       "CompALTA-MTA".Static_60 := 2;
   END_IF;
END_REGION

REGION Network 12
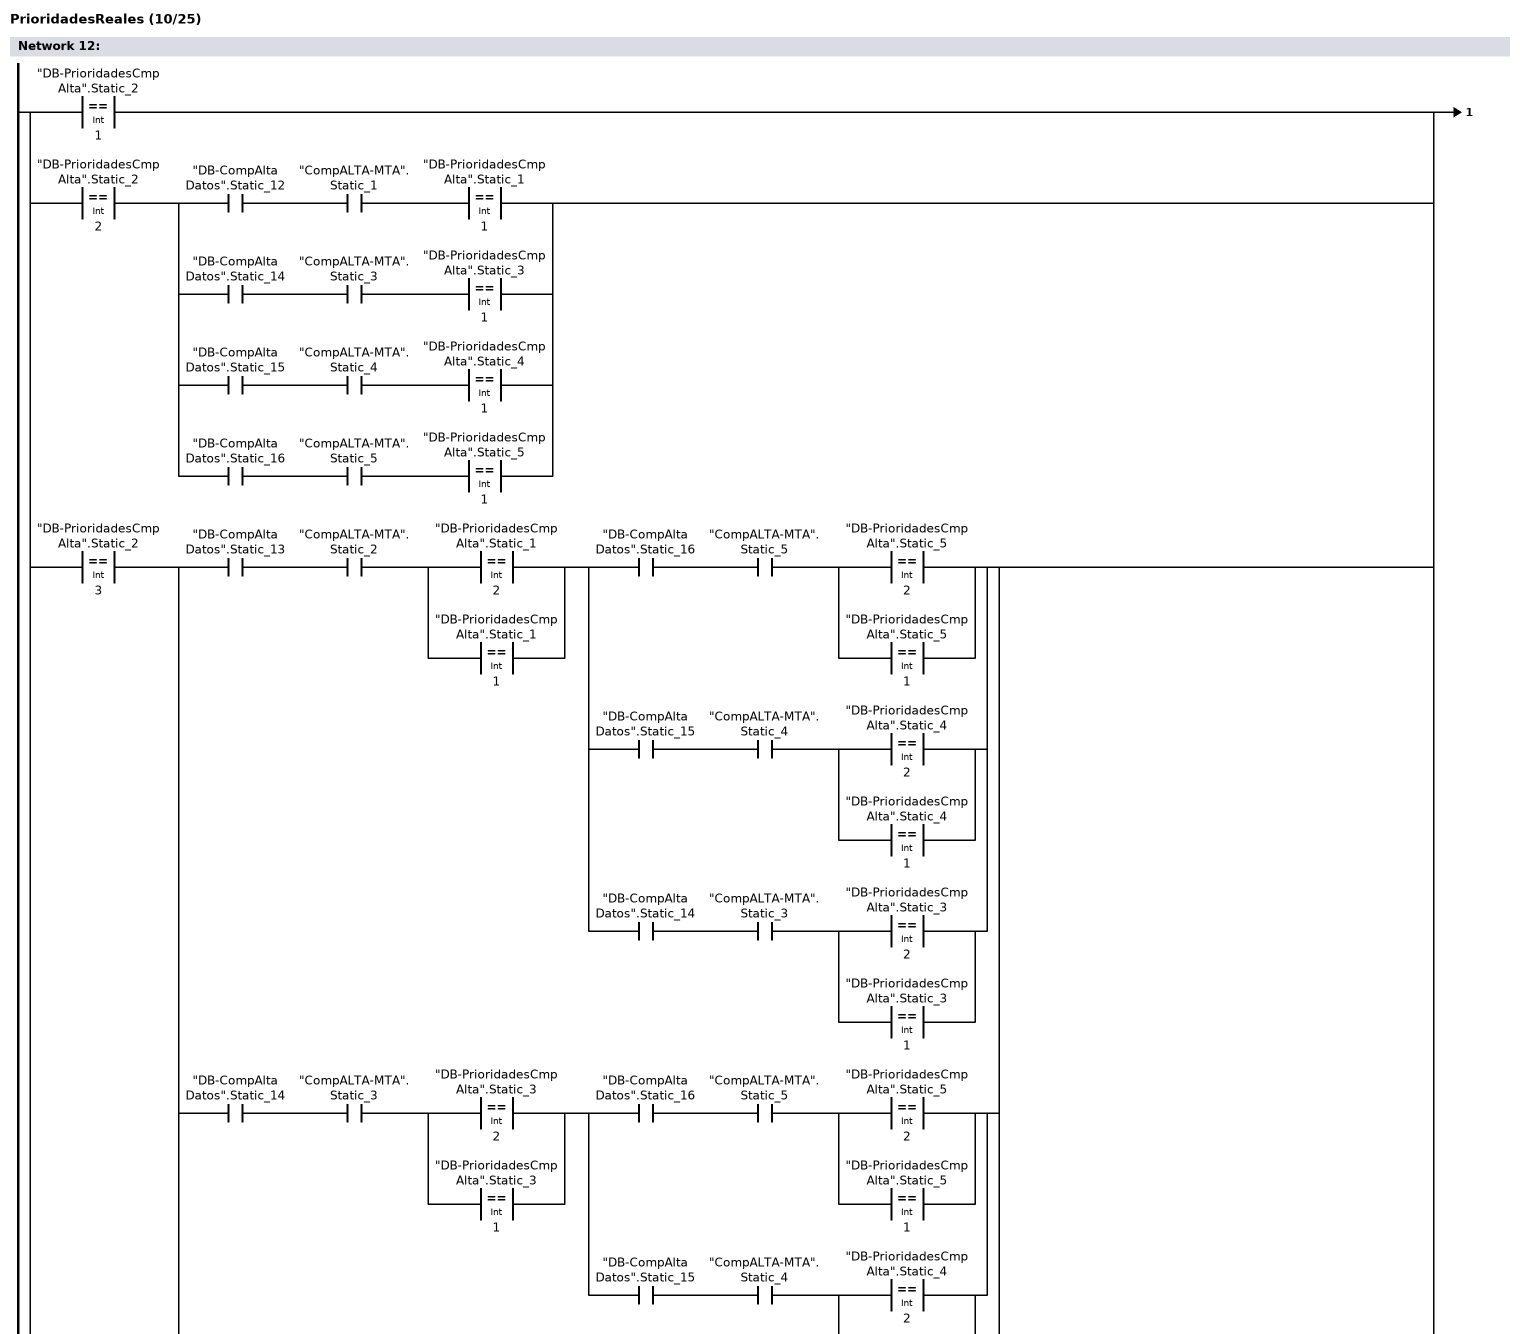
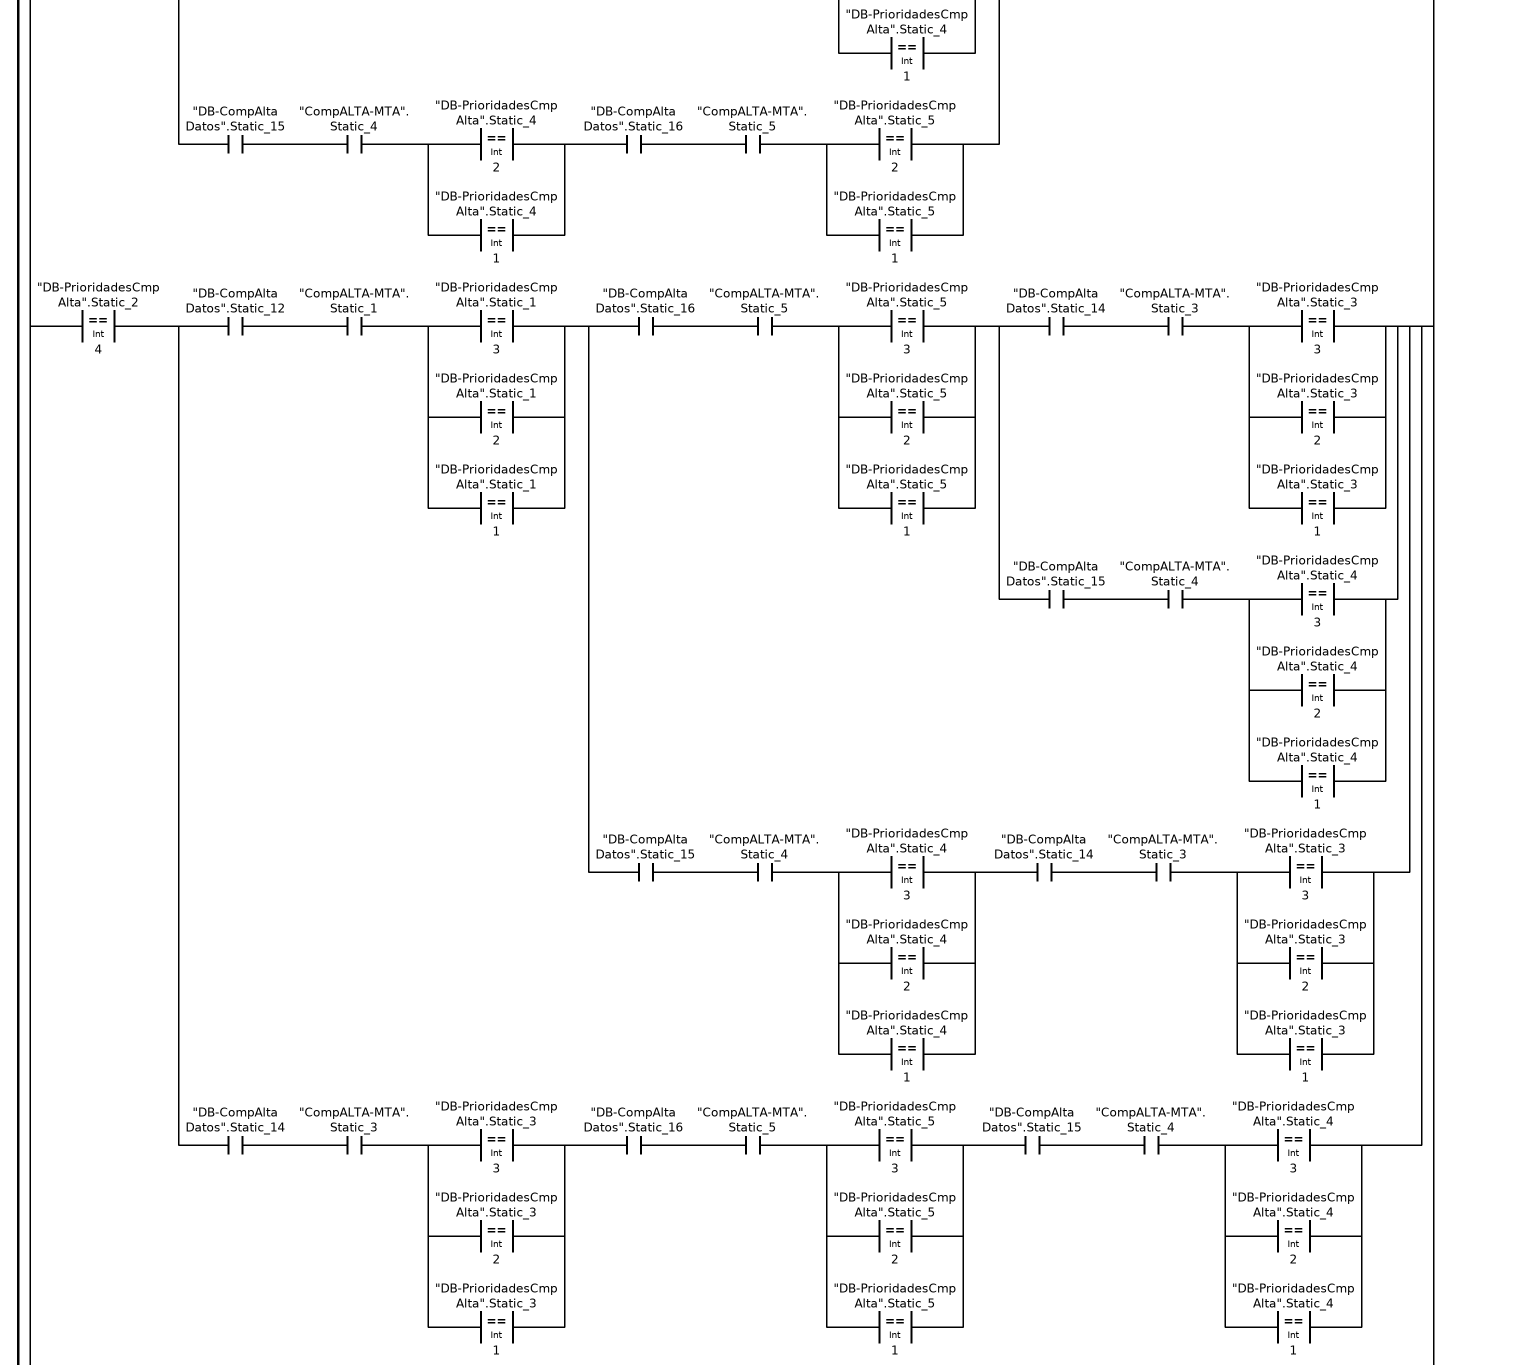
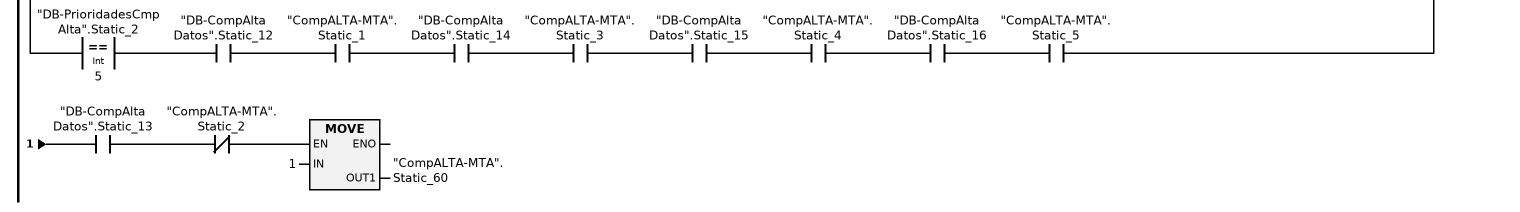
   IF (("DB-PrioridadesCmpAlta".Static_2 = 1) OR (("DB-PrioridadesCmpAlta".Static_2 = 2) AND (("DB-CompAltaDatos".Static_12 AND "CompALTA-MTA".Static_1 AND ("DB-PrioridadesCmpAlta".Static_1 = 1)) OR ("DB-CompAltaDatos".Static_14 AND "CompALTA-MTA".Static_3 AND ("DB-PrioridadesCmpAlta".Static_3 = 1)) OR ("DB-CompAltaDatos".Static_15 AND "CompALTA-MTA".Static_4 AND ("DB-PrioridadesCmpAlta".Static_4 = 1)) OR ("DB-CompAltaDatos".Static_16 AND "CompALTA-MTA".Static_5 AND ("DB-PrioridadesCmpAlta".Static_5 = 1)))) OR (("DB-PrioridadesCmpAlta".Static_2 = 3) AND (("DB-CompAltaDatos".Static_13 AND "CompALTA-MTA".Static_2 AND (("DB-PrioridadesCmpAlta".Static_1 = 2) OR ("DB-PrioridadesCmpAlta".Static_1 = 1)) AND (("DB-CompAltaDatos".Static_16 AND "CompALTA-MTA".Static_5 AND (("DB-PrioridadesCmpAlta".Static_5 = 2) OR ("DB-PrioridadesCmpAlta".Static_5 = 1))) OR ("DB-CompAltaDatos".Static_15 AND "CompALTA-MTA".Static_4 AND (("DB-PrioridadesCmpAlta".Static_4 = 2) OR ("DB-PrioridadesCmpAlta".Static_4 = 1))) OR ("DB-CompAltaDatos".Static_14 AND "CompALTA-MTA".Static_3 AND (("DB-PrioridadesCmpAlta".Static_3 = 2) OR ("DB-PrioridadesCmpAlta".Static_3 = 1))))) OR ("DB-CompAltaDatos".Static_14 AND "CompALTA-MTA".Static_3 AND (("DB-PrioridadesCmpAlta".Static_3 = 2) OR ("DB-PrioridadesCmpAlta".Static_3 = 1)) AND (("DB-CompAltaDatos".Static_16 AND "CompALTA-MTA".Static_5 AND (("DB-PrioridadesCmpAlta".Static_5 = 2) OR ("DB-PrioridadesCmpAlta".Static_5 = 1))) OR ("DB-CompAltaDatos".Static_15 AND "CompALTA-MTA".Static_4 AND (("DB-PrioridadesCmpAlta".Static_4 = 2) OR ("DB-PrioridadesCmpAlta".Static_4 = 1))))) OR ("DB-CompAltaDatos".Static_15 AND "CompALTA-MTA".Static_4 AND (("DB-PrioridadesCmpAlta".Static_4 = 2) OR ("DB-PrioridadesCmpAlta".Static_4 = 1)) AND "DB-CompAltaDatos".Static_16 AND "CompALTA-MTA".Static_5 AND (("DB-PrioridadesCmpAlta".Static_5 = 2) OR ("DB-PrioridadesCmpAlta".Static_5 = 1))))) OR (("DB-PrioridadesCmpAlta".Static_2 = 4) AND (("DB-CompAltaDatos".Static_12 AND "CompALTA-MTA".Static_1 AND (("DB-PrioridadesCmpAlta".Static_1 = 3) OR ("DB-PrioridadesCmpAlta".Static_1 = 2) OR ("DB-PrioridadesCmpAlta".Static_1 = 1)) AND (("DB-CompAltaDatos".Static_16 AND "CompALTA-MTA".Static_5 AND (("DB-PrioridadesCmpAlta".Static_5 = 3) OR ("DB-PrioridadesCmpAlta".Static_5 = 2) OR ("DB-PrioridadesCmpAlta".Static_5 = 1)) AND (("DB-CompAltaDatos".Static_14 AND "CompALTA-MTA".Static_3 AND (("DB-PrioridadesCmpAlta".Static_3 = 3) OR ("DB-PrioridadesCmpAlta".Static_3 = 2) OR ("DB-PrioridadesCmpAlta".Static_3 = 1))) OR ("DB-CompAltaDatos".Static_15 AND "CompALTA-MTA".Static_4 AND (("DB-PrioridadesCmpAlta".Static_4 = 3) OR ("DB-PrioridadesCmpAlta".Static_4 = 2) OR ("DB-PrioridadesCmpAlta".Static_4 = 1))))) OR ("DB-CompAltaDatos".Static_15 AND "CompALTA-MTA".Static_4 AND (("DB-PrioridadesCmpAlta".Static_4 = 3) OR ("DB-PrioridadesCmpAlta".Static_4 = 2) OR ("DB-PrioridadesCmpAlta".Static_4 = 1)) AND "DB-CompAltaDatos".Static_14 AND "CompALTA-MTA".Static_3 AND (("DB-PrioridadesCmpAlta".Static_3 = 3) OR ("DB-PrioridadesCmpAlta".Static_3 = 2) OR ("DB-PrioridadesCmpAlta".Static_3 = 1))))) OR ("DB-CompAltaDatos".Static_14 AND "CompALTA-MTA".Static_3 AND (("DB-PrioridadesCmpAlta".Static_3 = 3) OR ("DB-PrioridadesCmpAlta".Static_3 = 2) OR ("DB-PrioridadesCmpAlta".Static_3 = 1)) AND "DB-CompAltaDatos".Static_16 AND "CompALTA-MTA".Static_5 AND (("DB-PrioridadesCmpAlta".Static_5 = 3) OR ("DB-PrioridadesCmpAlta".Static_5 = 2) OR ("DB-PrioridadesCmpAlta".Static_5 = 1)) AND "DB-CompAltaDatos".Static_15 AND "CompALTA-MTA".Static_4 AND (("DB-PrioridadesCmpAlta".Static_4 = 3) OR ("DB-PrioridadesCmpAlta".Static_4 = 2) OR ("DB-PrioridadesCmpAlta".Static_4 = 1))))) OR (("DB-PrioridadesCmpAlta".Static_2 = 5) AND "DB-CompAltaDatos".Static_12 AND "CompALTA-MTA".Static_1 AND "DB-CompAltaDatos".Static_14 AND "CompALTA-MTA".Static_3 AND "DB-CompAltaDatos".Static_15 AND "CompALTA-MTA".Static_4 AND "DB-CompAltaDatos".Static_16 AND "CompALTA-MTA".Static_5)) AND "DB-CompAltaDatos".Static_13 AND NOT "CompALTA-MTA".Static_2 THEN
       "CompALTA-MTA".Static_60 := 1;
   END_IF;
END_REGION

REGION Network 15
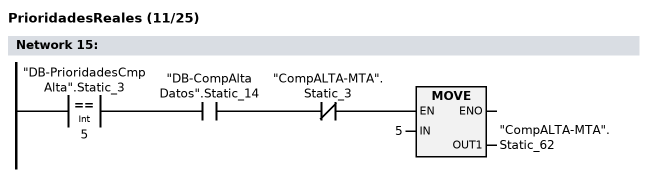
   RUNG wire#powerrail
      { S7_Templates := "SrcType := Int" } EQ_Contact(in1 := "DB-PrioridadesCmpAlta".Static_3, in2 := 5)
      Contact( "DB-CompAltaDatos".Static_14 )
      I_Contact( "CompALTA-MTA".Static_3 )
      { S7_GenerateENO := "TRUE" } Move(in := 5, out1 => "CompALTA-MTA".Static_62)
   END_RUNG
   // the same network as SCL:
   IF ("DB-PrioridadesCmpAlta".Static_3 = 5) AND "DB-CompAltaDatos".Static_14 AND NOT "CompALTA-MTA".Static_3 THEN
       "CompALTA-MTA".Static_62 := 5;
   END_IF;
END_REGION

REGION Network 16
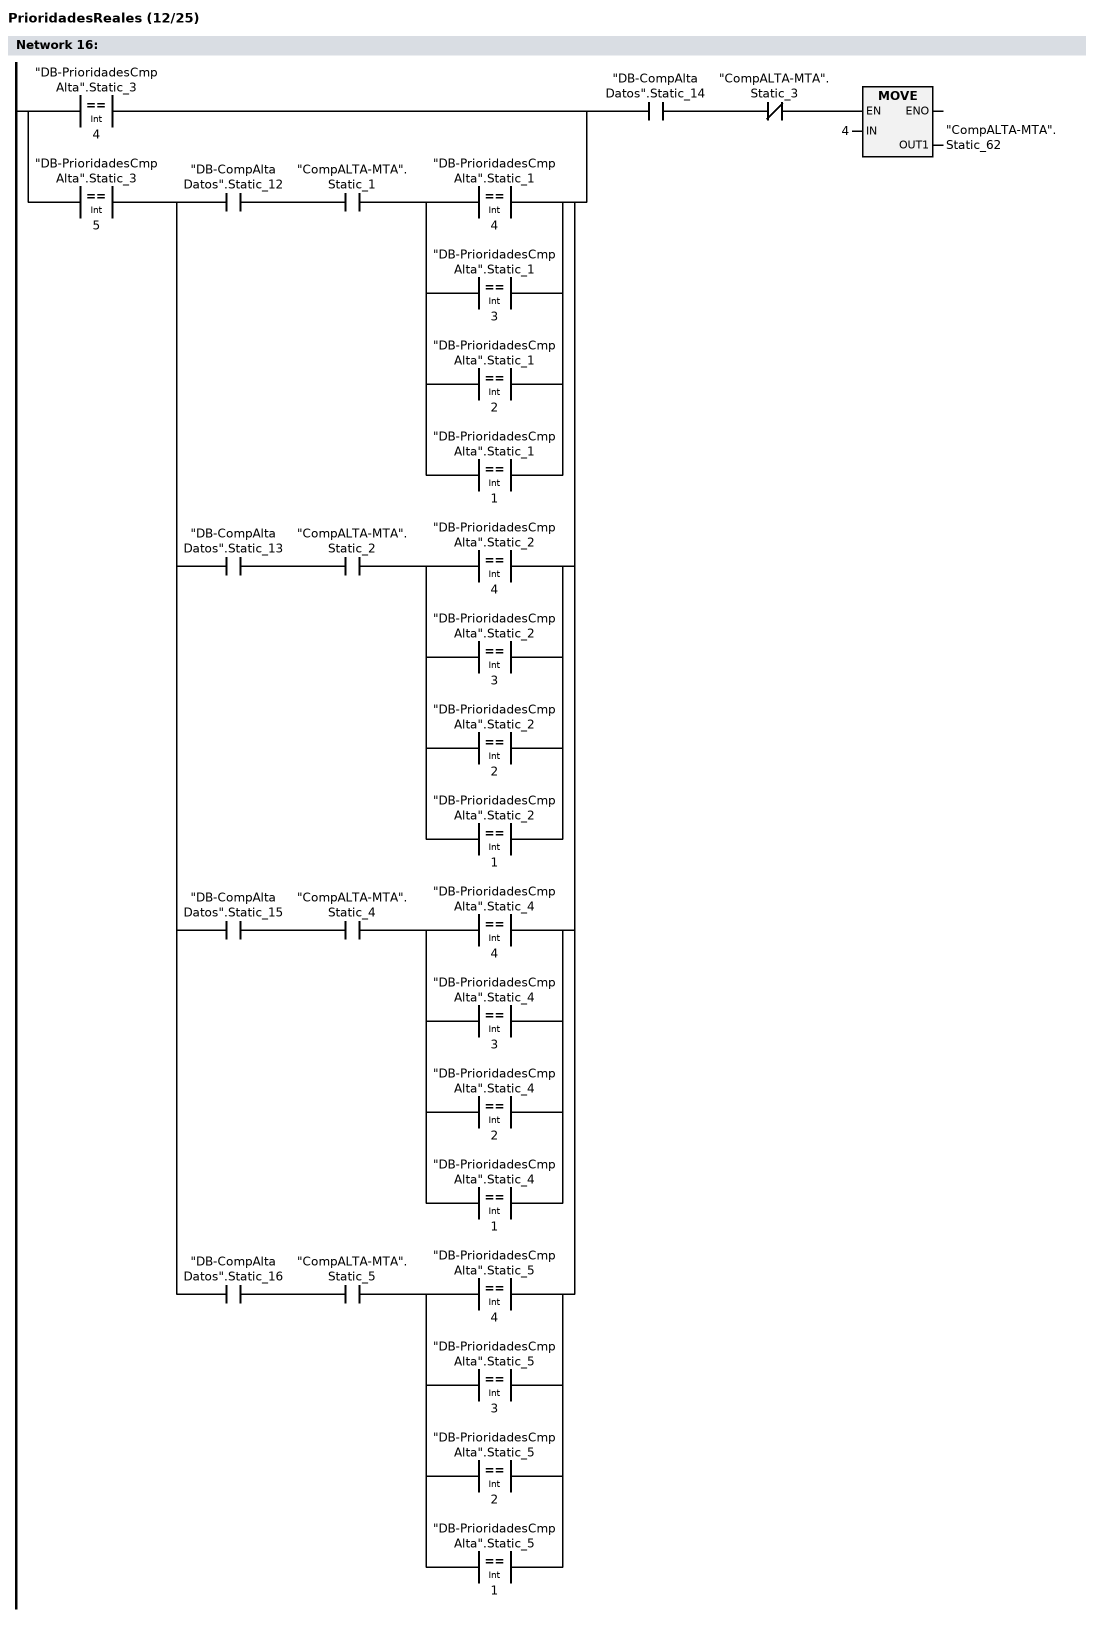
   IF (("DB-PrioridadesCmpAlta".Static_3 = 4) OR (("DB-PrioridadesCmpAlta".Static_3 = 5) AND (("DB-CompAltaDatos".Static_12 AND "CompALTA-MTA".Static_1 AND (("DB-PrioridadesCmpAlta".Static_1 = 4) OR ("DB-PrioridadesCmpAlta".Static_1 = 3) OR ("DB-PrioridadesCmpAlta".Static_1 = 2) OR ("DB-PrioridadesCmpAlta".Static_1 = 1))) OR ("DB-CompAltaDatos".Static_13 AND "CompALTA-MTA".Static_2 AND (("DB-PrioridadesCmpAlta".Static_2 = 4) OR ("DB-PrioridadesCmpAlta".Static_2 = 3) OR ("DB-PrioridadesCmpAlta".Static_2 = 2) OR ("DB-PrioridadesCmpAlta".Static_2 = 1))) OR ("DB-CompAltaDatos".Static_15 AND "CompALTA-MTA".Static_4 AND (("DB-PrioridadesCmpAlta".Static_4 = 4) OR ("DB-PrioridadesCmpAlta".Static_4 = 3) OR ("DB-PrioridadesCmpAlta".Static_4 = 2) OR ("DB-PrioridadesCmpAlta".Static_4 = 1))) OR ("DB-CompAltaDatos".Static_16 AND "CompALTA-MTA".Static_5 AND (("DB-PrioridadesCmpAlta".Static_5 = 4) OR ("DB-PrioridadesCmpAlta".Static_5 = 3) OR ("DB-PrioridadesCmpAlta".Static_5 = 2) OR ("DB-PrioridadesCmpAlta".Static_5 = 1)))))) AND "DB-CompAltaDatos".Static_14 AND NOT "CompALTA-MTA".Static_3 THEN
       "CompALTA-MTA".Static_62 := 4;
   END_IF;
END_REGION

REGION Network 17
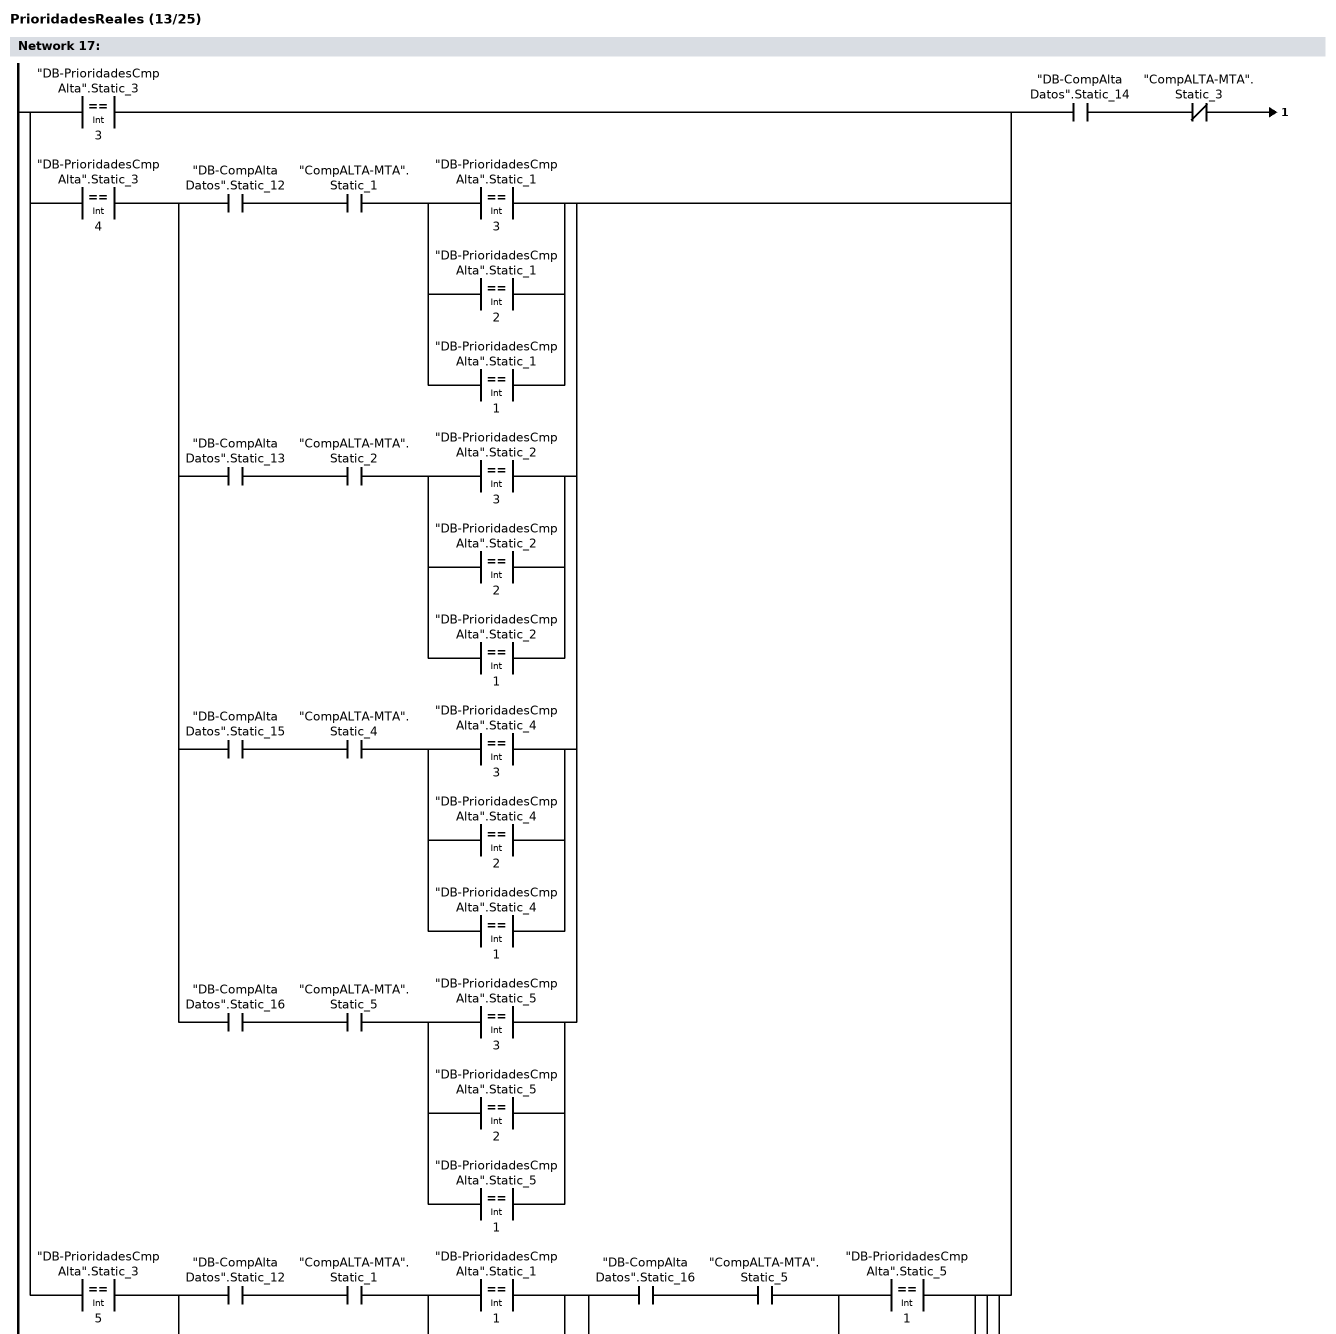
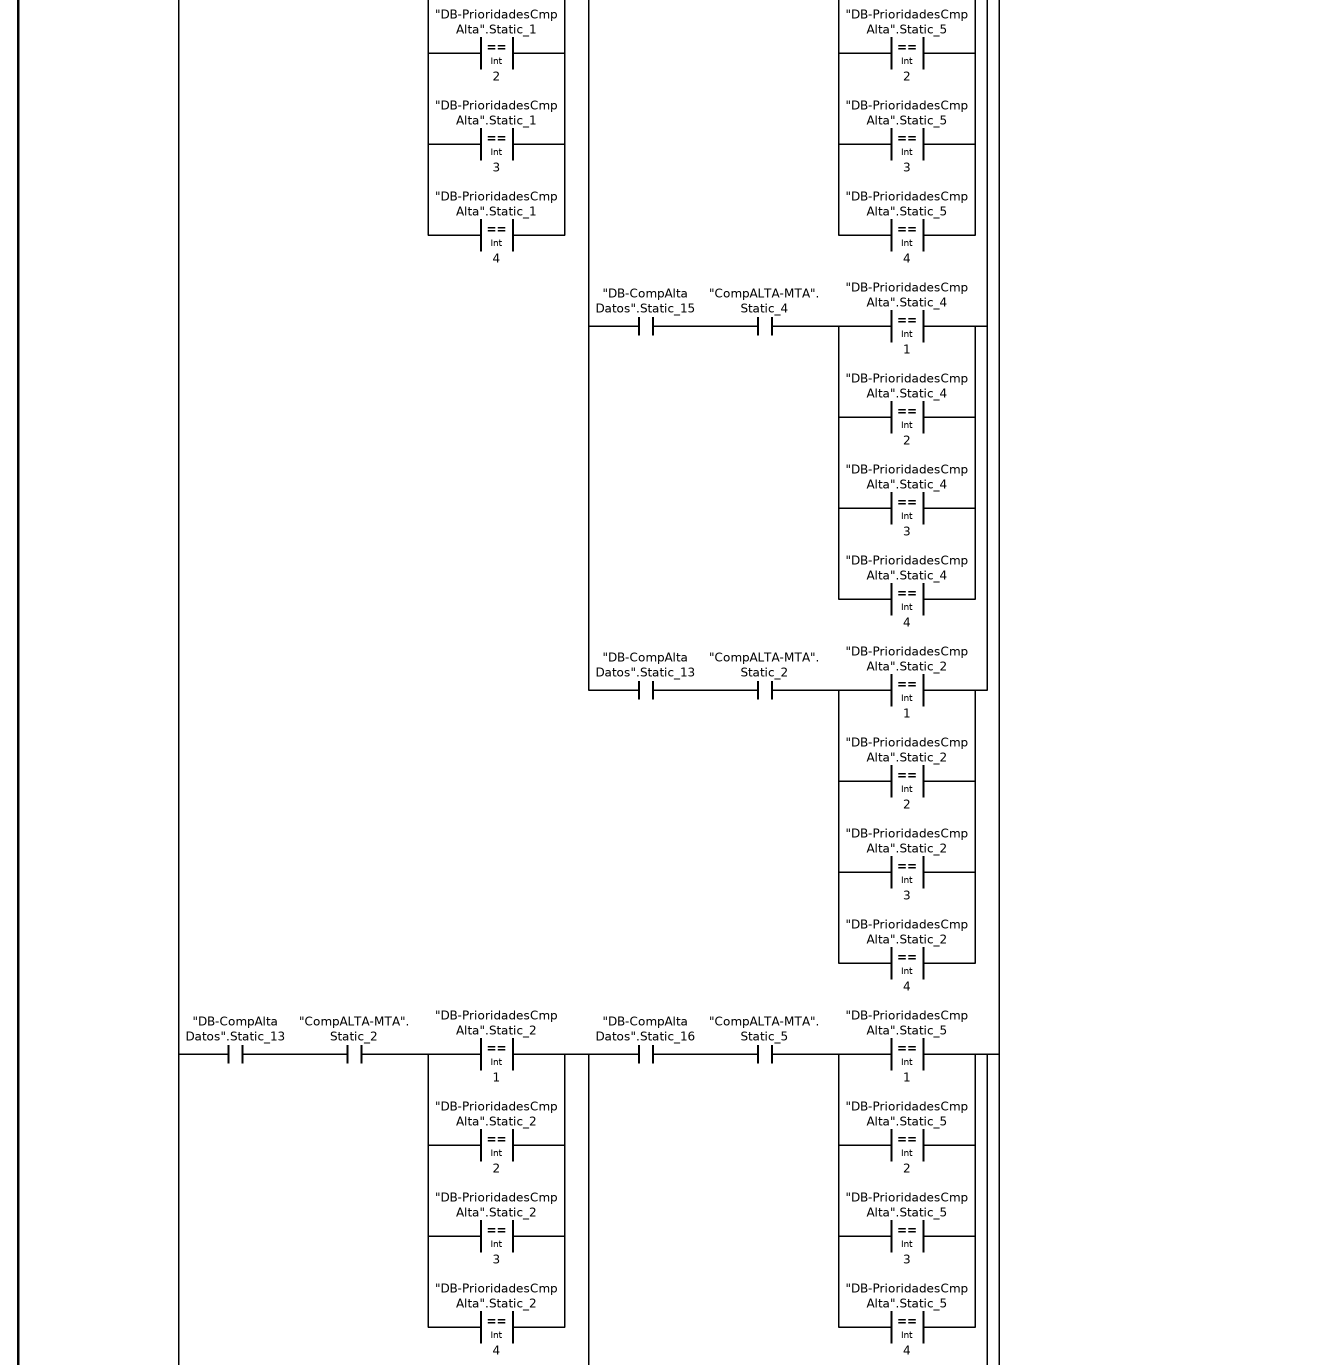
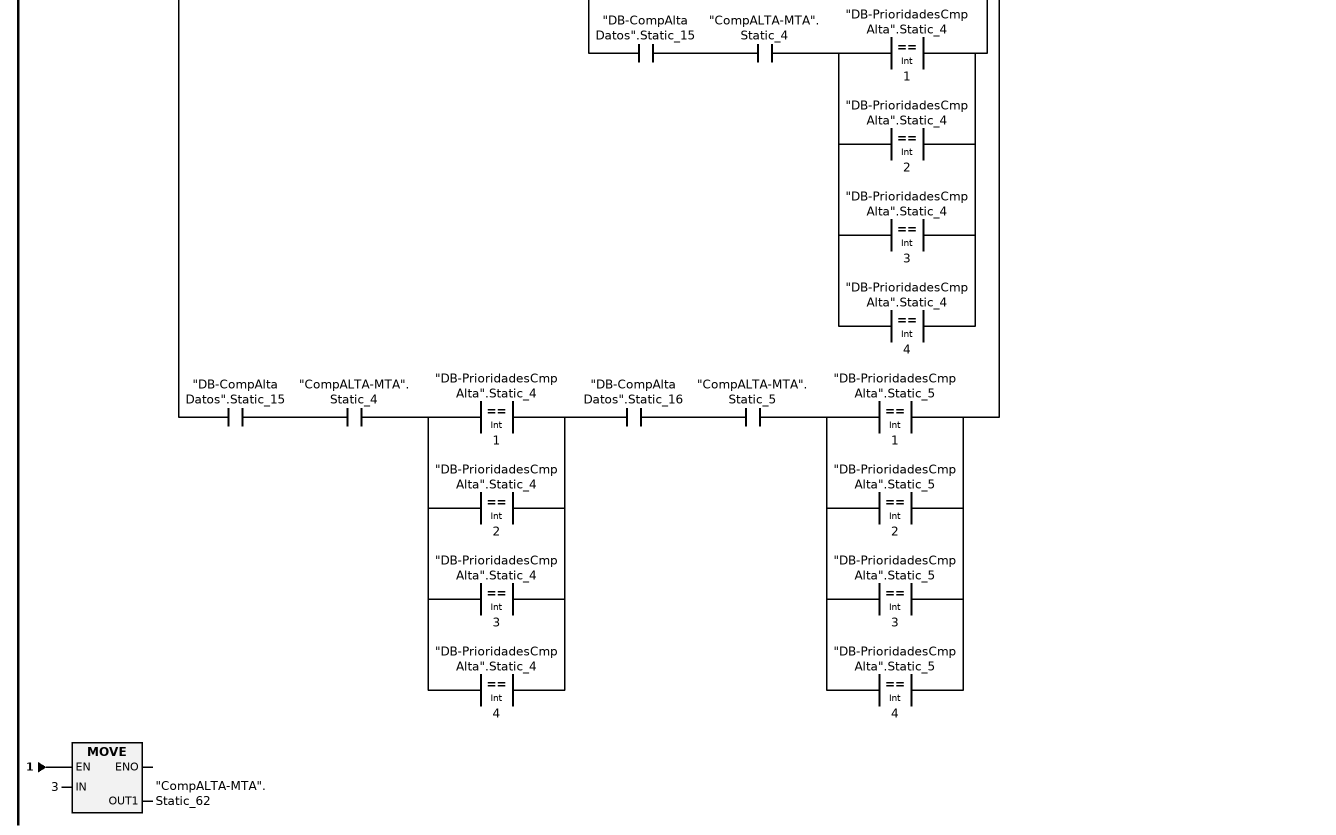
   IF (("DB-PrioridadesCmpAlta".Static_3 = 3) OR (("DB-PrioridadesCmpAlta".Static_3 = 4) AND (("DB-CompAltaDatos".Static_12 AND "CompALTA-MTA".Static_1 AND (("DB-PrioridadesCmpAlta".Static_1 = 3) OR ("DB-PrioridadesCmpAlta".Static_1 = 2) OR ("DB-PrioridadesCmpAlta".Static_1 = 1))) OR ("DB-CompAltaDatos".Static_13 AND "CompALTA-MTA".Static_2 AND (("DB-PrioridadesCmpAlta".Static_2 = 3) OR ("DB-PrioridadesCmpAlta".Static_2 = 2) OR ("DB-PrioridadesCmpAlta".Static_2 = 1))) OR ("DB-CompAltaDatos".Static_15 AND "CompALTA-MTA".Static_4 AND (("DB-PrioridadesCmpAlta".Static_4 = 3) OR ("DB-PrioridadesCmpAlta".Static_4 = 2) OR ("DB-PrioridadesCmpAlta".Static_4 = 1))) OR ("DB-CompAltaDatos".Static_16 AND "CompALTA-MTA".Static_5 AND (("DB-PrioridadesCmpAlta".Static_5 = 3) OR ("DB-PrioridadesCmpAlta".Static_5 = 2) OR ("DB-PrioridadesCmpAlta".Static_5 = 1))))) OR (("DB-PrioridadesCmpAlta".Static_3 = 5) AND (("DB-CompAltaDatos".Static_12 AND "CompALTA-MTA".Static_1 AND (("DB-PrioridadesCmpAlta".Static_1 = 1) OR ("DB-PrioridadesCmpAlta".Static_1 = 2) OR ("DB-PrioridadesCmpAlta".Static_1 = 3) OR ("DB-PrioridadesCmpAlta".Static_1 = 4)) AND (("DB-CompAltaDatos".Static_16 AND "CompALTA-MTA".Static_5 AND (("DB-PrioridadesCmpAlta".Static_5 = 1) OR ("DB-PrioridadesCmpAlta".Static_5 = 2) OR ("DB-PrioridadesCmpAlta".Static_5 = 3) OR ("DB-PrioridadesCmpAlta".Static_5 = 4))) OR ("DB-CompAltaDatos".Static_15 AND "CompALTA-MTA".Static_4 AND (("DB-PrioridadesCmpAlta".Static_4 = 1) OR ("DB-PrioridadesCmpAlta".Static_4 = 2) OR ("DB-PrioridadesCmpAlta".Static_4 = 3) OR ("DB-PrioridadesCmpAlta".Static_4 = 4))) OR ("DB-CompAltaDatos".Static_13 AND "CompALTA-MTA".Static_2 AND (("DB-PrioridadesCmpAlta".Static_2 = 1) OR ("DB-PrioridadesCmpAlta".Static_2 = 2) OR ("DB-PrioridadesCmpAlta".Static_2 = 3) OR ("DB-PrioridadesCmpAlta".Static_2 = 4))))) OR ("DB-CompAltaDatos".Static_13 AND "CompALTA-MTA".Static_2 AND (("DB-PrioridadesCmpAlta".Static_2 = 1) OR ("DB-PrioridadesCmpAlta".Static_2 = 2) OR ("DB-PrioridadesCmpAlta".Static_2 = 3) OR ("DB-PrioridadesCmpAlta".Static_2 = 4)) AND (("DB-CompAltaDatos".Static_16 AND "CompALTA-MTA".Static_5 AND (("DB-PrioridadesCmpAlta".Static_5 = 1) OR ("DB-PrioridadesCmpAlta".Static_5 = 2) OR ("DB-PrioridadesCmpAlta".Static_5 = 3) OR ("DB-PrioridadesCmpAlta".Static_5 = 4))) OR ("DB-CompAltaDatos".Static_15 AND "CompALTA-MTA".Static_4 AND (("DB-PrioridadesCmpAlta".Static_4 = 1) OR ("DB-PrioridadesCmpAlta".Static_4 = 2) OR ("DB-PrioridadesCmpAlta".Static_4 = 3) OR ("DB-PrioridadesCmpAlta".Static_4 = 4))))) OR ("DB-CompAltaDatos".Static_15 AND "CompALTA-MTA".Static_4 AND (("DB-PrioridadesCmpAlta".Static_4 = 1) OR ("DB-PrioridadesCmpAlta".Static_4 = 2) OR ("DB-PrioridadesCmpAlta".Static_4 = 3) OR ("DB-PrioridadesCmpAlta".Static_4 = 4)) AND "DB-CompAltaDatos".Static_16 AND "CompALTA-MTA".Static_5 AND (("DB-PrioridadesCmpAlta".Static_5 = 1) OR ("DB-PrioridadesCmpAlta".Static_5 = 2) OR ("DB-PrioridadesCmpAlta".Static_5 = 3) OR ("DB-PrioridadesCmpAlta".Static_5 = 4)))))) AND "DB-CompAltaDatos".Static_14 AND NOT "CompALTA-MTA".Static_3 THEN
       "CompALTA-MTA".Static_62 := 3;
   END_IF;
END_REGION

REGION Network 18
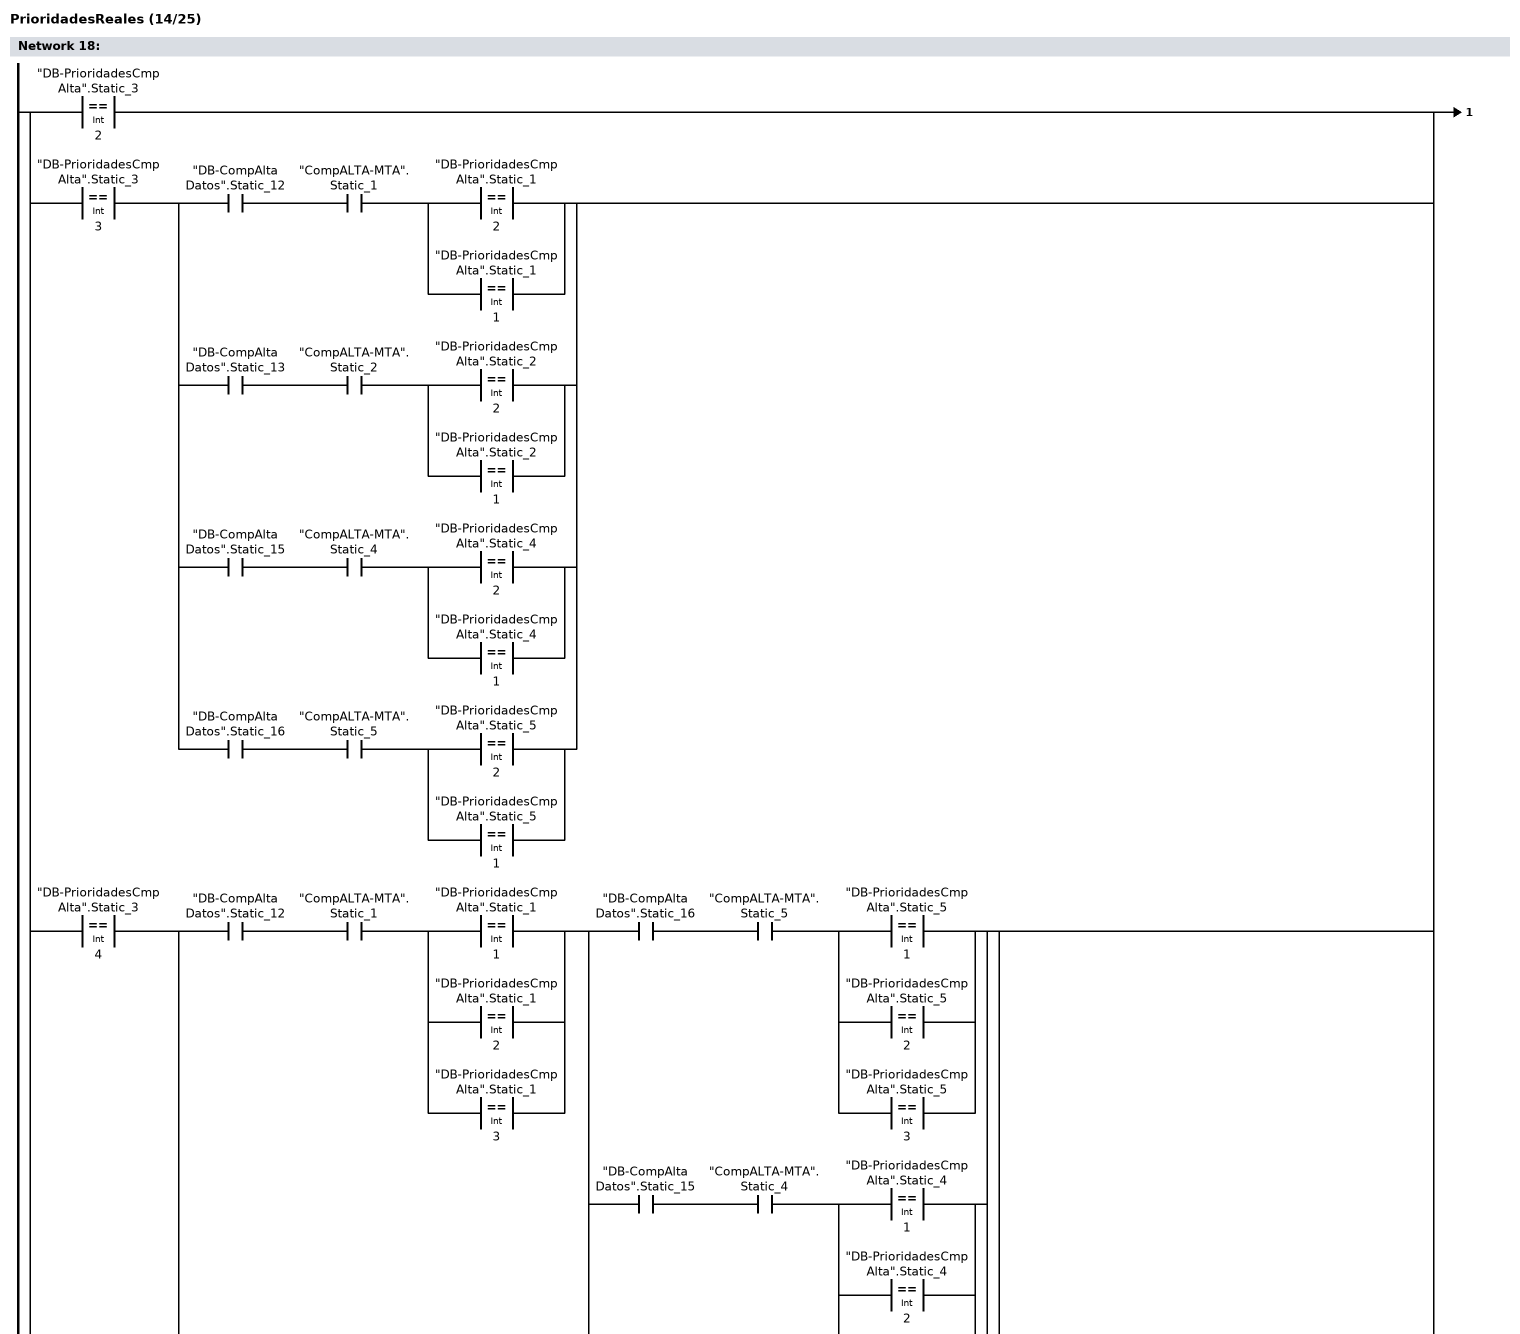
